// TIA Portal project "e009004v440" (V15.1) (continued)
   40: 'Reserva', class Reserva, trigger "DB_OP.DEF03" bit 15
   87: 'Falla al cerrar pinza posicionadora: Comprobar Sensores 29S4 y 29S5 + Electroválvula 43Y8 / FORMAGE : DEF MOUVEMENT FERMETURE PINCE 43Y8 : vérifier 29S4 29S5', class Fallos Pinza, trigger "DB_OP.DEF06" bit 14
   19: 'Falla térmica en freno de motor ajuste de ancho en etapa de Formado: Comprobar estado de Guardamotor Q09 / DF_QF9_1', class Fallos Formado, trigger "DB_OP.DEF02" bit 10
   68: 'Falla al subir araña: Comprobar sensores 25S7 y 25S8, y electroválvula 41Y3 / Falla al subir Araña: Comprobar Sensores 25S7 y 25S8 + Electroválvula 41Y3 / PREHENSEUR : DEF MOUVEMENT MONTEE 41Y3 : vérifier 25S7 25S8', class Fallos Araña, trigger "DB_OP.DEF05" bit 11
   71: 'Reserva', class Reserva, trigger "DB_OP.DEF05" bit 14
   21: 'Falla de excursión en Ajuste de ancho de Perfiladores: Comprobar 29S6, 29S7 + Encóder correspondiente / DEFAUT MOP PROFILEUSE : vérifier 29S6 29S7 ou codeur DP15', class Fallos Perfiladores, trigger "DB_OP.DEF02" bit 12
   67: 'Falla al bajar Araña: Comprobar Sensores 25S7 y 25S8 + Electroválvula 41Y2 / PREHENSEUR : DEF MOUVEMENT DESCENTE 41Y2 : vérifier 25S7 25S8', class Fallos Araña, trigger "DB_OP.DEF05" bit 10
   5: 'Falla en Variador Transporte Rolos: Comprobar estado de Variador VAR03 / Variateur OK Convoyeur Magasin', class Fallos Rolos, trigger "DB_OP.DEF01" bit 12
   24: 'Reserva', class Reserva, trigger "DB_OP.DEF02" bit 15
   95: 'Incoherencia en lectura de sensores 26S6 (Araña Arriba) y 26S7 (Araña Abajo) Soluciones Posibles: - Revise que el estado de ambos sensores sea correcto. - Revise el cableado de ambos sensores y asegúrese de que las señales llegan al panel observando los estados de los mismos desde el esquemático del PANEL / Falla al avanzar intercambiador de Almacenes: Comprobar Sensores 26S6 y 26S7 + Contactor KM01.1 / CHARGEMENT : DEF MOUVEMENT AVANCE MAGASIN : vérifier 26S6 26S7', class Fallos Almacenes, trigger "DB_OP.DEF06" bit 6
   101: 'Falla al subir Herramienta de Formado: Comprobar Sensores 28S5 y 28S6 + Relé 43K4 / FORMAGE : DEF MOUVEMENT MONTEE OUTIL 43K4 : vérifier 28S5 28S6', class Fallos Formado, trigger "DB_OP.DEF07" bit 12
   20: 'Falla en presión hidráulica en freno Perfiladores: Comprobar Sensor 23S4 / DEFAUT PRESSION HYDRAULIQUE FREIN PROFILEUSE : Vérifier 23S4', class Fallos Perfiladores, trigger "DB_OP.DEF02" bit 11
   50: 'Falla en Plegador 1 al intentar realizar plegado: Comprobar Sensores 31S7 y 31S8 + Relé 45K5 / PLIEUSE 1 : DEF MOUVEMENT AVANCE PLIAGE 45K5 : vérifier 31S7 et 31S8', class Fallos Plegadora, trigger "DB_OP.DEF04" bit 9
   111: 'Reserva', class Reserva, trigger "DB_OP.DEF07" bit 6
   65: 'Falla al transladar Araña (Avance): Comprobar Sensores 26S2 y 26S3 + Contactor KM02.1 / PREHENSEUR : DEF MOUVEMENT AVANCE KM02_1 : vérifier 26S2 26S3', class Fallos Araña, trigger "DB_OP.DEF05" bit 8
   53: 'Falla en Plegador 2 al intentar activar fijación: Comprobar Sensores 35S1 y 35S2 + Relé 47K1 / PLIEUSE 1 : DEF MOUVEMENT AVANCE BRIDAGE 45K3 : vérifier 31S5 et 31S6', class Fallos Plegadora, trigger "DB_OP.DEF04" bit 12
   109: 'Reserva', class Reserva, trigger "DB_OP.DEF07" bit 4
   39: 'Reserva', class Reserva, trigger "DB_OP.DEF03" bit 14
   56: 'Falla en Plegador 2 al intentar bajar primera extensión de prensa: Comprobar Sensores 35S7 y 35S8 + Relé 46K7 / PLIEUSE 2 : DEF MOUVEMENT AVANCE V2 47K7 : vérifier 35S7 et 35S8', class Fallos Plegadora, trigger "DB_OP.DEF04" bit 15
   54: 'Falla en Plegador 2 al intentar realizar plegado: Comprobar Sensores 35S3 y 35S4 + Relé 47K3 / PLIEUSE 1 : DEF MOUVEMENT AVANCE PLIAGE 45K5 : vérifier 31S7 et 31S8', class Fallos Plegadora, trigger "DB_OP.DEF04" bit 13
   108: 'Reserva', class Reserva, trigger "DB_OP.DEF07" bit 3
   86: 'Falla al bajar Bloqueador de Avance en etapa formador: Comprobar Sensores 29S1 y 29S2 + Electroválvula 43Y5 / FORMAGE : DEF MOUVEMENT DESCENTE BUTEE 43Y5 : vérifier 29S1 29S2', class Fallos Formado, trigger "DB_OP.DEF06" bit 13
   93: 'Falla al bajar Herramienta de Formado: Comprobar Sensores 28S5 y 28S6 + Relé 43K3 / FORMAGE : DEF MOUVEMENT DESCENTE OUTIL 43K3 : vérifier 28S5 28S6', class Fallos Formado, trigger "DB_OP.DEF06" bit 4
   34: 'Falla al bajar pinza en Plegadora: Comprobar Sensores 30S3 y 30S4 + Electroválvula 44Y3 / PLIEUSE : DEF MOUVEMENT DESCENTE PINCE 44Y3 : vérifier 30S3 et 30S4', class Fallos Plegadora, trigger "DB_OP.DEF03" bit 9
   27: 'Falla presión de Aire: Comprobar estado del Presostato 23S7 / DEFAUT AIR', class Fallos Generales, trigger "DB_OP.DEF02" bit 2
   115: 'Reserva', class Reserva, trigger "DB_OP.DEF08" bit 10
   97: 'Falla al retroceder martillo de herramienta 1 en Formador: Comprobar Sensores 27S5 y 27S6 + Relé 42K4 / FORMAGE : DEF MOUVEMENT RECUL MARTEAU OUTIL 1 42K4 : vérifier 27S5 27S6', class Fallos Formado, trigger "DB_OP.DEF07" bit 8
   88: 'Reserva', class Reserva, trigger "DB_OP.DEF06" bit 15
   57: 'Falla en Plegador 1 al intentar desactivar fijación: Comprobar Sensores 31S5 y 31S6 + Relé 45K4 / PLIEUSE 1 : DEF MOUVEMENT RECUL BRIDAGE 45K4 : vérifier 31S5 et 31S6', class Fallos Plegadora, trigger "DB_OP.DEF04" bit 0
   26: 'Falla de seguridad: Comprobar seguridades y relé de seguridad KAU1 / ATTENTE MISE EN SERVICE', class Fallos Generales, trigger "DB_OP.DEF02" bit 1
   18: 'Falla térmica en motor grupo hidráulico Plegadora: Comprobar estado de Guardamotor QM013.1 / DF_QM013_1 PLIEUSE : Moteur Groupe HYdraulique', class Fallos Plegadora, trigger "DB_OP.DEF02" bit 9
   36: 'Falla al activar alineacion X de Pieza en Plegadora: Comprobar Sensores 21S5, 21S6, 36S1 y 36S2 + Relé 46K5 / PLIEUSE : DEF MOUVEMENT TAQUAGE X 46K5 : vérifier 21S5 21S6 36S1 36S2', class Fallos Plegadora, trigger "DB_OP.DEF03" bit 11
   7: 'Falla en etapa de Potencia de variadores Perfiladores: Comprobar el estado de U13.2, U13.9, U13.12, U13.15 y U13.17 en Tablero T02 / DF_QM04 PROFILEUSE : Moteur 1,2,3 ou 4', class Fallos Perfiladores, trigger "DB_OP.DEF01" bit 14
   25: 'Falla alimentación de Entradas: Comprrobar estado de Térmica Q6 / ATTENTE MISE SOUS TENSION', class Fallos Generales, trigger "DB_OP.DEF02" bit 0
   104: 'Reserva', class Reserva, trigger "DB_OP.DEF07" bit 0
   96: 'Reserva', class Reserva, trigger "DB_OP.DEF06" bit 7
   77: 'Falla en Plegador 1 al intentar subir segunda extensión de prensa: Comprobar Sensores 32S5 y 32S6 + Relé 46K3 / PLIEUSE 1 : DEF MOUVEMENT AVANCE V3 46K3 : vérifier 32S5 32S6', class Fallos Plegadora, trigger "DB_OP.DEF05" bit 4
   8: 'Falla presente en CU Plegadores: Compruebe estado de CPU10', class Fallos Plegadora, trigger "DB_OP.DEF01" bit 15
   78: 'Falla en Plegador 2 al intentar subir segunda extensión de prensa: Comprobar Sensores 35S7 y 35S8 + Relé 48K1 / PLIEUSE 1 : DEF MOUVEMENT AVANCE V3 46K3 : vérifier 32S5 32S6', class Fallos Plegadora, trigger "DB_OP.DEF05" bit 5
   17: 'Falla límite de Seguridad en Plegador 2: Compruebe Sensor límite de carrera correspondiente / DF_VAR12 :PLIEUSE 2 : ServoVariateur OK', class Fallos Plegadora, trigger "DB_OP.DEF02" bit 8
   75: 'Reserva', class Reserva, trigger "DB_OP.DEF05" bit 2
   106: 'Reserva', class Reserva, trigger "DB_OP.DEF07" bit 1
   1: 'Falla térmica en motor refrigeración de grupo hidráulico Plegadora: Comprobar estado de Guardamotor QM013.2 / Moteur OK refroidisseur GH plieuse', class Fallos Perfiladores, trigger "DB_OP.DEF01" bit 8
   9: 'Falla de seguridad presente en CU Plegadores: Compruebe estado de CPU10', class Fallos Plegadora, trigger "DB_OP.DEF01" bit 0
   84: 'Reserva', class Reserva, trigger "DB_OP.DEF06" bit 11
   98: 'Falla al retroceder matriz de herramienta 1 en Formador: Comprobar Sensores 27S7 y 27S8 + Relé 42K6 / FORMAGE : DEF MOUVEMENT RECUL MATRICE OUTIL 1 42K6 : vérifier 27S7 27S8', class Fallos Formado, trigger "DB_OP.DEF07" bit 9
   92: 'Falla al avanzar matriz de herramienta 2 en Formador: Comprobar Sensores 28S3 y 28S4 + Relé 43K1 / FORMAGE : DEF MOUVEMENT AVANCE MATRICE OUTIL 2 43K1 : vérifier 28S3 28S4', class Fallos Formado, trigger "DB_OP.DEF06" bit 3
   99: 'Falla al retroceder martillo de herramienta 1 en Formador: Comprobar Sensores 28S1 y 28S2 + Relé 42K8 / FORMAGE : DEF MOUVEMENT RECUL MARTEAU OUTIL 2 42K8 : vérifier 28S1 28S2', class Fallos Formado, trigger "DB_OP.DEF07" bit 10
   120: 'Reserva', class Reserva, trigger "DB_OP.DEF08" bit 15
   16: 'Falla límite de Seguridad en Plegador 1: Compruebe Sensor límite de carrera correspondiente', class Fallos Plegadora, trigger "DB_OP.DEF01" bit 7
   59: 'Falla en Plegador 1 al intentar subir prensa: Comprobar Sensores 32S1 y 32S2 + Relé 45K8 / PLIEUSE 1 : DEF MOUVEMENT RECUL V1 45K8 : vérifier 32S1 et 32S2', class Fallos Plegadora, trigger "DB_OP.DEF04" bit 2
   42: 'Falla al subir pinza en Plegadora: Comprobar Sensores 30S3 y 30S4 + Electroválvula 44Y4 / PLIEUSE : DEF MOUVEMENT MONTEE PINCE 44Y4 : vérifier 30S3 et 30S4', class Fallos Plegadora, trigger "DB_OP.DEF03" bit 1
   11: 'Falla térmica en grupo hidraulico de freno Perfiladores: Comprobar estado de Guardamotor QM06 / DF_QM06 : PROFILEUSE : GH frein OK', class Fallos Perfiladores, trigger "DB_OP.DEF01" bit 2
   102: 'Falla al retroceder Descargador: Comprobar Sensores 31S2 y 31S3 + Relé 45K2 / DECHARGEMENT : DEF RECUL ESCAMOTEUR 45K2 : vérifier 31S2 31S3', class Fallos Descargador, trigger "DB_OP.DEF07" bit 13
   52: 'Falla en Plegador 1 al intentar subir primera extensión de prensa: Comprobar Sensores 32S3 y 32S4 + Relé 46K1', class Fallos Plegadora, trigger "DB_OP.DEF04" bit 11
   76: 'Reserva', class Reserva, trigger "DB_OP.DEF05" bit 3
   81: 'Falla al avanzar ajuste de formado: Comprobar Contactor KM09.1 + Encóder correspondiente / FORMAGE : DEF MOUVEMENT AVANCE MOP KM09_1 : vérifier codeur 2', class Fallos Cinta, trigger "DB_OP.DEF06" bit 8
   107: 'Reserva', class Reserva, trigger "DB_OP.DEF07" bit 2
   15: 'Falla Rectificador de variadores Plegadores: Comprobar estado de AL10', class Fallos Plegadora, trigger "DB_OP.DEF01" bit 6
   80: 'Falla en Plegador 2 al intentar bajar segunda extensión de prensa: Comprobar Sensores 35S7 y 35S8 + Relé 48K2 / PLIEUSE 1 : DEF MOUVEMENT AVANCE V3 46K3 : vérifier 32S5 32S6', class Fallos Plegadora, trigger "DB_OP.DEF05" bit 7
   47: 'Reserva', class Reserva, trigger "DB_OP.DEF03" bit 6
   43: 'Falla al cerrar pinza en Plegadora: Comprobar Sensores 30S5 y 30S6 + Electroválvula 44Y6 / PLIEUSE : DEF MOUVEMENT FERMETURE PINCE 44Y6 : vérifier 30S5 et 30S6', class Fallos Plegadora, trigger "DB_OP.DEF03" bit 2
   13: 'Falla en Variador Transporte Cinta: Comprobar estado de VAR08 / DF_VAR08 : CONVOYEUR 2 : Variateur OK', class Fallos Cinta, trigger "DB_OP.DEF01" bit 4
   45: 'Falla al desactivar alineacion Y de Pieza en Plegadora: Comprobar Sensores 23S6 y 36S4 + Relé 46K6', class Fallos Plegadora, trigger "DB_OP.DEF03" bit 4
   105: 'Reserva', class Reserva, trigger "DB_OP.DEF07" bit 15
   38: 'Falla al desactivar alineacion Y de Pieza en Plegadora: Comprobar Sensores 23S5, 23S6, 36S3 y 36S4 + Relé 46K6', class Fallos Plegadora, trigger "DB_OP.DEF03" bit 13
   31: 'Falla de Atasco de pieza en Perfilador: Compobar Sensores 36S13, 36S14, 36S15 y 36S16 / DEFAUT BOURRAGE PROFILEUSE', class Fallos Perfiladores, trigger "DB_OP.DEF02" bit 6
   72: 'Reserva', class Reserva, trigger "DB_OP.DEF05" bit 15
   89: 'Falla al avanzar martillo de herramienta 1 en Formador: Comprobar Sensores 27S5 y 27S6 + Relé 42K3 / FORMAGE : DEF MOUVEMENT AVANCE MARTEAU OUTIL 1 42K3 : vérifier 27S5 27S6', class Fallos Formado, trigger "DB_OP.DEF06" bit 0
   114: 'Reserva', class Reserva, trigger "DB_OP.DEF08" bit 9
   10: 'Falla térmica en bomba de lubricación de Perfiladores: Comprobar estado de Guardamotor QM05 / DF_QM05 : PROFILEUSE :Pompes lubrifications OK', class Fallos Perfiladores, trigger "DB_OP.DEF01" bit 1
   4: 'Falla en Variador Transporte de Araña: Comprobar estado de Variador VAR02 / Variateur OK Axe Prehenseur', class Fallos Araña, trigger "DB_OP.DEF01" bit 11
   110: 'Reserva', class Reserva, trigger "DB_OP.DEF07" bit 5
   73: 'Falla al transladar Araña (Retroceder): Comprobar Sensores 26S2 y 26S3, y Contactor KM02.2 / PREHENSEUR : DEF MOUVEMENT RECUL KM02_2 : vérifier 26S2 26S3', class Fallos Araña, trigger "DB_OP.DEF05" bit 0
   44: 'Falla al desactivar alineacion X de Pieza en Plegadora: Comprobar Sensores 36S2 y 21S6 + Relé 46K5 / PLIEUSE : DEF MOUVEMENT TAQUAGE X 46K5 : vérifier 21S5 21S6 36S1 36S2', class Fallos Plegadora, trigger "DB_OP.DEF03" bit 3
   118: 'Reserva', class Reserva, trigger "DB_OP.DEF08" bit 13
   94: 'Falla al avanzar Descargador: Comprobar Sensores 31S2 y 31S3 + Relé 45K1 / DECHARGEMENT : DEF AVANCE ESCAMOTEUR 45K1 : vérifier 31S2 31S3', class Fallos Descargador, trigger "DB_OP.DEF06" bit 5
   58: 'Falla en Plegador 1 al intentar desactivar orden de plegado: Comprobar Sensores 31S7 y 31S8 + Relé 45K6 / PLIEUSE 1 : DEF MOUVEMENT RECUL PLIAGE 45K6 : vérifier 31S7 et 31S8', class Fallos Plegadora, trigger "DB_OP.DEF04" bit 1
   63: 'Falla en Plegador 2 al intentar subir prensa: Comprobar Sensores 35S5 y 35S6 + Relé 47K6 / PLIEUSE 1 : DEF MOUVEMENT RECUL V1 45K8 : vérifier 32S1 et 32S2', class Fallos Plegadora, trigger "DB_OP.DEF04" bit 6
   119: 'Reserva', class Reserva, trigger "DB_OP.DEF08" bit 14
   60: 'Falla en Plegador 1 al intentar bajar primera extensión de prensa: Comprobar Sensores 32S3 y 32S4 + Relé 46K2', class Fallos Plegadora, trigger "DB_OP.DEF04" bit 3
   23: 'Falla Seguridad de Perímetro: Comprobar Seguridad de puertas y tablero CPI / DF_RES01', class Fallos Generales, trigger "DB_OP.DEF02" bit 14
   32: 'Reserva / DF_RES01', class Reserva, trigger "DB_OP.DEF02" bit 7
   22: 'Falla de excursión en Ajuste de ancho de Formado: Comprobar 28S7, 28S8 + Encóder correspondiente / DEFAUT MOP CONVOYEUR2 : vérifier 28S7 28S8 ou codeur DP16', class Fallos Formado, trigger "DB_OP.DEF02" bit 13
   79: 'Falla en Plegador 1 al intentar bajar segunda extensión de prensa: Comprobar Sensores 32S5 y 32S6 + Relé 46K3 / PLIEUSE 2 : DEF MOUVEMENT AVANCE V3 48K1 : vérifier 36S7 36S8', class Fallos Plegadora, trigger "DB_OP.DEF05" bit 6

text list "SelecciónPlegadora": 0 'Sin selección'; 1 'Plegador 1'; 2 'Plegador 2'; 3 'Tenaza'

text list "Modo": 0 'Detenido / ARRET'; 1 'Modo Manual / MANUEL'; 2 'Modo Automático / AUTO'; 3 'En Ciclo / CYCLE'; 4 'Finalizando Ciclo / FIN CYCLE'

text list "RC1": 0 '00: Sin selección / 00: ACQUITTEMENT'; 1 '01: Intercambiador de almacenes - Avance / 01 : Avance Magasin (mag 1)'; 2 '02: Intercambiador de almacenes - Retroceso / 02 : Recul Magasin (mag 2)'; 11 '11: Transporte Araña - Avance / 11 : Préhenseur Avance'; 12 '12: Transporte Araña - Retroceso / 12 : Préhenseur Recul'; 13 '13: Araña - Bajar sobre Almacén 1 / 13 : Préhenseur Magasin 1'; 14 '14: Araña - Bajar sobre Almacén 2 / 14 : Préhenseur Magasin 2'; 15 '15: Araña - Bajar / 15 : Préhenseur Descente'; 16 '16: Araña - Subir / 16 : Préhenseur Montée'; 20 '20: Tulipas de Araña - Aire en todas ON / 20 :Flambage 1 à 3 Avance'; 21 '21: Tulipas de Araña - Aire en todas OFF / 21: Flambage 1 à 3 Recul'; 22 '22: Tulipas de Araña - Aire en Grupo 1 ON / 22 : Flambage 1 Avance'; 23 '23: Tulipas de Araña - Aire en Grupo 1 OFF / 23 : Flambage 1 Recul'; 24 '24: Tulipas de Araña - Aire en Grupo 2 ON / 24 : Flambage 2 Avance'; 25 '25: Tulipas de Araña - Aire en Grupo 2 OFF / 25 : Flambage 2 Recul'; 26 '26: Tulipas de Araña - Aire en Grupo 3 ON / 26 : Flambage 3 Avance'; 27 '27: Tulipas de Araña - Aire en Grupo 3 OFF / 27 : Flambage 3 Recul'; 30 '30: Tulipas de Araña - Vacío en Todas ON / 30 :Aspiration 1 à 3 Avance'; 31 '31: Tulipas de Araña - Vacío en Todas OFF / 31: Aspiration 1 à 3 Recul'; 32 '32: Tulipas de Araña - Vacío en Grupo 1 ON / 32 : Aspiration 1 Avance'; 33 '33: Tulipas de Araña - Vacío en Grupo 1 OFF / 33 : Aspiration 1 Recul'; 34 '34 : Tulipas de Araña - Vacío en Grupo 2 ON / 34 : Aspiration 2 Avance'; 35 '35: Tulipas de Araña - Vacío en Grupo 2 OFF / 35 : Aspiration 2 Recul'; 36 '36: Tulipas de Araña - Vacío en Grupo 3 ON / 36 : Aspiration 3 Avance'; 37 '37: Tulipas de Araña - Vacío en Grupo 3 OFF / 37 : Aspiration 3 Recul'; 41 '41: Transporte Rolos - Avance / 41 avance Convoyeur 1'; 42 '42: Transporte Rolos - Retroceso / 42 Recul Convoyeur 1'; 51 '51: Ajuste de profundidad Perfiladores - Hacia Consigna / 51 : MOP Profileuse Consigne'; 52 '52: Ajuste de profundidad Perfiladores - Cerrar / 52 : Avance MOP Profileuse'; 53 '53: Ajuste de profundidad Perfiladores - Abrir / 53 : Recul MOP Profileuse'; 54 '54: Ajuste de profundidad Perfiladores - Freno / 54 : Frein MOP profileuse'; 55 '55: Perfiladores - Retroceso / 55 : Avance Profileuse'; 56 '56: Perfiladores - Avance / 56 : Recul Profileuse'

text list "RC2": 0 '00: Sin Selección / 00: ACQUITTEMENT'; 1 '01: Plegadora - Avance Tenaza / 01:Pince: Avance'; 2 '02: Plegadora - Retroceso Tenaza / 02:Pince: Recul'; 3 '03: Plegadora - Bajar Tenaza / 03:Pince: Descente'; 4 '04: Plegadora - Subir Tenaza / 04:Pince: Montée'; 5 '05: Plegadora - Abrir Tenaza / 05:Pince: ouverture'; 6 '06: Plegadora - Cerrar Tenaza / 06:Pince: Fermeture'; 7 '07: Plegadora - Alineación X / 07:taquage X'; 8 '08: Plegadora - Alineación Y / 08:taquage Y'; 9 '09: Plegadora - Subir Cepillos / 09: brosse'; 10 '10: Plegador 1 - Bloquear Prensa / 10:PLIEUSE 1: bridage Avance'; 11 '11: Plegador 1 - Desbloquear Prensa / 11:PLIEUSE 1: bridage Recul'; 12 '12: Plegador 1 - Bajar Prensa / 12:PLIEUSE 1: V1 Avance'; 13 '13: Plegador 1 - Subir Prensa / 13:PLIEUSE 1: V1 Recul'; 14 '14: Plegador 1 - Bajar Extension Prensa 1 / 14:PLIEUSE 1: V2 Avance'; 15 '15: Plegador 1 - Subir Extension Prensa 1 / 15:PLIEUSE 1: V2 Recul'; 16 '16: Plegador 1 - Bajar Extension Prensa 2 / 16:PLIEUSE 1: V3 Avance'; 17 '17: Plegador 1 - Subir Extension Prensa 2 / 17:PLIEUSE 1: V3 Recul'; 18 '18: Plegador 1 - Subir / 18:PLIEUSE 1: Montée'; 19 '19: Plegador 1 - Bajar / 19:PLIEUSE 1: Descente'; 20 '20: Plegador 2 - Bloquear Prensa / 20:PLIEUSE 2: bridage Avance'; 21 '21: Plegador 2 - Desbloquear Prensa / 21:PLIEUSE 2: bridage Recul'; 22 '22: Plegador 2 - Bajar Prensa / 22:PLIEUSE 2: V1 Avance'; 23 '23: Plegador 2 - Subir Prensa / 23:PLIEUSE 2: V1 Recul'; 24 '24: Plegador 2 - Bajar Extension Prensa 1 / 22:PLIEUSE 2: V1 Avance'; 25 '25: Plegador 2 - Subir Extension Prensa 1 / 23:PLIEUSE 2: V1 Recul'; 26 '26: Plegador 2 - Bajar Extension Prensa 2 / 26:PLIEUSE 2: V3 Avance'; 27 '27: Plegador 2 - Subir Extension Prensa 2 / 27:PLIEUSE 2: V3 Recul'; 28 '28: Plegador 2 - Subir / 28:PLIEUSE 2: Montée'; 29 '29: Plegador 2 - Bajar / 29:PLIEUSE 2: Descente'; 31 '31: Pinza - Avance / 31 : Avance Pince'; 32 '32: Pinza - Retroceso / 32 : Recul Pince'; 33 '33: Pinza - Abrir / 33: Ouverture Pince'; 34 '34: Pinza - Cerrar / 34: Fermeture Pince'; 35 '35: Formador - Subir Tope / 35: Montée Butée'; 36 '36: Formador - Bajar Tope / 36: Descente Butée'; 37 '37: Formador - Ajuste de profundidad - Hacia Consigna / 37: Position Consigne'; 38 '38: Formador - Ajuste de profundidad - Avance / 38: Rapproche ( - )'; 39 '39: Formador - Ajuste de profundidad - Retroceso / 39: Ecartement ( + )'; 40 '40: Formador - Bajar Herramientas / 40: Descente Ensemble'; 41 '41: Formador - Subir Herramientas / 41: Montée Ensemble'; 42 '42: Formador - Herramienta 1 - Martillo ON / 42: MARTEAU : Avance Outil 1'; 43 '43: Formador - Herramienta 1 - Martillo OFF / 43: MARTEAU : Recul Outil 1'; 44 '44: Formador - Herramienta 1 - Matriz ON / 44: MATRICE : Avance Outil 1'; 45 '45: Formador - Herramienta 1 - Matriz OFF / 45: MATRICE : Recul Outil 1'; 46 '46: Formador - Herramienta 2 - Martillo ON / 46: MARTEAU : Avance Outil 2'; 47 '47: Formador - Herramienta 2 - Martillo OFF / 47: MARTEAU : Recul Outil 2'; 48 '48: Formador - Herramienta 2 - Matriz ON / 48: MATRICE : Avance Outil 2'; 49 '49: Formador - Herramienta 2 - Matriz OFF / 49: MATRICE : Recul Outil 2'; 61 '61: Plegador 1 - Avance (apertura) / 61: PLIEUSE 1 : Ecartement +'; 62 '62: Plegador 1 - Retroceso (cierre) / 62: PLIEUSE 1 : Rapproche -'; 65 '65: Plegador 2 - Avance (apertura) / 65: PLIEUSE 2 : Ecartement +'; 66 '66: Plegador 2 - Retroceso (cierre) / 66: PLIEUSE 2 : Rapproche -'; 70 '70: Descargador - Avance / 70: Avance Escamoteur'; 71 '71: Descargador - Retroceso / 71: Recul Escamoteur'; 91 '91: Transporte Cinta - Avance / 91: Avance Convoyeur 2'; 92 '92: Transporte Cinta - Retroceso / 92: Recul Convoyeur 2'

text list "Warnings": 0 'Sin Warnings'; 1 'Reconocimiento de Fallas solo es posible en Modo Manual'; 2 'No es posible intercambiar almacenes si la Araña no está completamente arriba'; 4 ''; 8 'Los plegadores no pueden desplazarse si sus prensas no estan completamente abiertas'; 16 'Los plegados solo son posibles con las prensas abajo'; 32 'Para poder bloquear los plegadores es becesario que las prensas estén abajo'; 64 'Solo es posible accionar las herramientas si el formador está abajo'; 128 ''; 254 ''; 512 ''; 1024 ''; 2048 ''; 4096 ''

text list "Estados_PL": 0 'Detenido'; 512 'Esperando Pieza'; 1024 'Ingresando Pieza'; 2048 'Posicionando Plegadores para Primer Plegado'; 4096 'Realizando Primer Plegado'; 8192 'Realizando Segundo Plegado'; 16384 'Entregando Pieza'; 2 'Alineando Pieza'; 4 'Posicionando Plegadores para Segundo Plegado'; 8 'Posicionando Plegadores para Entrega de Pieza'; 16 'Posicionando Plegadores para Espera'

text list "Estados_F": 128 'Detenido'; 512 'Esperando'; 1024 'Formando Pieza en Esquina 1 con Herramienta 1'; 2048 'Formando Pieza en Esquina 1 con Herramienta 2'; 4096 'Formando Pieza en Esquina 2 con Herramienta 1'; 8192 'Formando Pieza en Esquina 2 con Herramienta 2'; 16384 'Entregando Pieza'; -32768 'Posicionando Pieza en Esquina 1 con Herramienta 1'; 1 'Posicionando Pieza en Esquina 1 con Herramienta 2'; 2 'Posicionando Pieza en Esquina 2 con Herramienta 1'; 4 'Posicionando Pieza en Esquina 2 con Herramienta 2'; 8 'Posicionando Pieza para Entrega'; 16 'Posicionando Pinza para Recepción de Pieza'

text list "Transiciones_PL": 0 'Condición de avance: Sin pieza en Plegadora'; 16 'Condición de avance: Posición de Espera alcanzada'; 512 'Condición de avance: Nueva Pieza en Plegadora'; 2 'Condición de avance: Alineadores Activos'; 2048 'Condición de avance: Posición de Plegado de Patas alcanzada'; 4 'Condición de avance: Posición de Plegado de Techo alcanzada'; 8 'Condición de avance: Posición de Entrega alcanzada'; 1024 'Condición de avance: Tenaza Plegadora adentro (Abierta)'; 4096 'Condición de avance: Plegado de Patas Activo'; 8192 'Condición de avance: Plegado de Techo Activo'; 16384 'Condición de avance: Pieza entregada a Descargador'

text list "Transiciones_F": 128 'Condición de avance: Sin Pieza en Pinza'; 512 'Condición de avance: Nueva Pieza en Final de Cinta'; 1024 'Condición de avance: Formado con Herramienta 1 Listo'; 2048 'Condición de avance: Formado con Herramienta 2 Listo'; 4096 'Condición de avance: Formado con Herramienta 1 Listo'; 8192 'Condición de avance: Formado con Herramienta 2 Listo'; 16384 'Condición de avance: Pieza entregada a Plegadora'; -32768 'Condición de avance: Posición de E1H1 alcanzada'; 1 'Condición de avance: Posición de E1H2 alcanzada'; 2 'Condición de avance: Posición de E2H1 alcanzada'; 4 'Condición de avance: Posición de E2H2 alcanzada'; 8 'Condición de avance: Posición de Entrega alcanzada'; 16 'Condición de avance: Posición de Recepción alcanzada'

text list "Proveedor": 0 ''; 1 'A'; 2 'B'; 3 'C'; 4 'D'; 5 'E'; 6 'F'

graphic list "General - Araña": 0..1 'Araña 1 G'; 1 'Araña 2_1'

graphic list "General - Almacén": 0..1 'Almacen 1 G'; 1 'Almacen 2_1'

graphic list "General - Rolos": 0..1 'Rolos 1 G'; 1 'Rolos 2_3'

graphic list "General - Perfiladores": 0..1 'Perfiladores 1 G'; 1 'Perfiladores 2_1'

graphic list "General - Cinta": 0..1 'Cinta G'; 1 'Cinta 2_1'

graphic list "General - Pinza": 0..1 'Pinza G'; 1 'Pinza 2_1'

graphic list "General - Formador": 0..1 'F1_G'; 1 'F1R'

graphic list "General - Plegadora": 0..1 'Plegador 1 G'; 1 'Plegador 2_1'

graphic list "General - Descargador": 0..1 'Descargador G'; 1 'Descargador 2_1'

graphic list "Intercambiador": 0..1 'ALM 2_1'; 1 'ALM 1'

graphic list "Grupo 3 - Plegadora": 0 'Pleg'; 1 'Pleg2'

graphic list "Grupo 3 - Descargador": 0..1 'Desc G'; 1 'Desc2'

graphic list "Grupo 3 - Pinza1": 0..1 'P2_G'; 1 'P2R'

graphic list "Pleg3": 1 'PLEG3b'; 2..3 'pleg_1'

graphic list "Grupo 1 - Rolos": 1 'Rolos 2 G'; 1 'Rolos 2b'

graphic list "Grupo 1 - Araña": 1 'Araña3b'; 2..3 'Araña3 G'

graphic list "Grupo 1 - Almacén A": 1 'ALM 2 G'; 2..3 'ALM 1 G'

graphic list "Grupo 1 - Almacén B": 1 'ALM 2b'; 2..3 'ALM 1b_1'

graphic list "Grupo 2 - Perfilador": 1 'PERFIb'; 2..3 'PERFI G'

graphic list "Grupo 2 - Cinta": 1 'CINb'; 2..3 'CIN G'

graphic list "Grupo 2 - Formador": 1 'Piqb'; 2..3 'Piq_1'

graphic list "Formador": 1 'F1R'; 2..3 'F1_G'

graphic list "Araña": 1 'Araña4b'; 2..3 'Araña4C'

graphic list "Rolos": 1 'Rolos 3b'; 2..3 'Rolos 3 G'

graphic list "GeneralBase": 0 'Base G'; 1 'BaseRoja'

graphic list "Estado": 0 'PilotLight_Round_GN_Off_256c'; 1 'PilotLight_Round_GN_On_256c'

graphic list "CheckBox": 0 'outline_check_box_outline_blank_black_18dp'; 1 'outline_check_box_black_18dp'

graphic list "CheckBox_Neg": 1 'outline_check_box_outline_blank_black_18dp'; 0 'outline_check_box_black_18dp'

graphic list "Pleg3_1": 1 'PLEG3b'; 2..3 'PLEG3_1'

graphic list "Grupo 3 - Pinza1_1": 0..1 'P2'; 1 'P2R'

graphic list "Formador_1": 1 'F2R'; 2..3 'F2C'

graphic list "Formador_2": 1 'F2R'; 2..3 'F2C'

recipe "Pieza": A <- "Receta\Recetas.A", B <- "Receta\Recetas.B", C <- "Receta\Recetas.C", D <- "Receta\Recetas.D", F1 <- "Receta\Recetas.F1", F2 <- "Receta\Recetas.F2", F3 <- "Receta\Recetas.F3", F4 <- "Receta\Recetas.F4", PL1_1 <- "Receta\Recetas.PL1_1", PL1_2 <- "Receta\Recetas.PL1_2", PL2_1 <- "Receta\Recetas.PL2_1", PL2_2 <- "Receta\Recetas.PL2_2"

screen "HabAlarmas9" 1280x768, template "Template"
   TextField "Campo de texto_1" at 117,85 size 37x18; Text '113 -'
   TextField "Campo de texto_2" at 117,129 size 37x18; Text '114 -'
   TextField "Campo de texto_3" at 117,173 size 37x18; Text '115 -'
   TextField "Campo de texto_4" at 117,217 size 367x18; Text '116 - Inconsistencia de Presencia de pieza en Transporte de Rolos'
   TextField "Campo de texto_5" at 117,261 size 37x18; Text '117 -'
   TextField "Campo de texto_6d" at 117,305 size 37x18; Text '118 -'
   TextField "Campo de texto_7" at 117,349 size 37x32; Text '119 -'
   TextField "Campo de texto_8" at 117,393 size 37x32; Text '120 -'
   TextField "Campo de texto_9" at 117,437 size 342x18; Text '121 - Inconsistencia de Presencia de pieza en en Descargador'
   Switch "Interruptor_1" at 48,77 size 59x33; TextOff 'SI'; TextOn 'NO'; CaptionText 'Switch'; PictureOff "Check"; PictureOn "UnCheck"
      ProcessValue <- "Desactivar_Falla113"
   Switch "Interruptor_2" at 48,121 size 59x33; TextOff 'SI'; TextOn 'NO'; CaptionText 'Switch'; PictureOff "Check"; PictureOn "UnCheck"
      ProcessValue <- "Desactivar_Falla114"
   Switch "Interruptor_3" at 48,165 size 59x33; TextOff 'SI'; TextOn 'NO'; CaptionText 'Switch'; PictureOff "Check"; PictureOn "UnCheck"
      ProcessValue <- "Desactivar_Falla115"
   Switch "Interruptor_4" at 48,209 size 59x33; TextOff 'SI'; TextOn 'NO'; CaptionText 'Switch'; PictureOff "Check"; PictureOn "UnCheck"
      ProcessValue <- "Desactivar_Falla116"
   Switch "Interruptor_5" at 48,253 size 59x33; TextOff 'SI'; TextOn 'NO'; CaptionText 'Switch'; PictureOff "Check"; PictureOn "UnCheck"
      ProcessValue <- "Desactivar_Falla117"
   Switch "Interruptor_6" at 48,297 size 59x33; TextOff 'SI'; TextOn 'NO'; CaptionText 'Switch'; PictureOff "Check"; PictureOn "UnCheck"
      ProcessValue <- "Desactivar_Falla118"
   Switch "Interruptor_7" at 48,341 size 59x33; TextOff 'SI'; TextOn 'NO'; CaptionText 'Switch'; PictureOff "Check"; PictureOn "UnCheck"
      ProcessValue <- "Desactivar_Falla119"
   Switch "Interruptor_8" at 48,385 size 59x33; TextOff 'SI'; TextOn 'NO'; CaptionText 'Switch'; PictureOff "Check"; PictureOn "UnCheck"
      ProcessValue <- "Desactivar_Falla120"
   Switch "Interruptor_9" at 48,429 size 59x33; TextOff 'SI'; TextOn 'NO'; CaptionText 'Switch'; PictureOff "Check"; PictureOn "UnCheck"
      ProcessValue <- "Desactivar_Falla121"
   TextField "Campo de texto_15" at 38,32 size 262x22; Text 'Configuración de habilitación de Alarmas'
   Button "Botón_2" at 1010,33 size 51x51; TextOff '<'
      on Click: ActivateScreen("HabAlarmas7", 0)
   Button "Botón_3" at 1202,33 size 51x51; TextOff '>'
   Circle "Círculo_2" at 24,87 size 12x12
      Appearance <- "Alarma 1"
   Circle "Círculo_3" at 25,131 size 12x12
      Appearance <- "Alarma 114"
   Circle "Círculo_4" at 25,175 size 12x12
      Appearance <- "Alarma 115"
   Circle "Círculo_5" at 24,87 size 12x12
      Appearance <- "Alarma 113"
   Circle "Círculo_6" at 25,219 size 12x12
      Appearance <- "Alarma 116"
   Circle "Círculo_7" at 25,263 size 12x12
      Appearance <- "Alarma 117"
   Circle "Círculo_8" at 25,307 size 12x12
      Appearance <- "Alarma 118"
   Circle "Círculo_9" at 25,351 size 12x12
      Appearance <- "Alarma 119"
   Circle "Círculo_10" at 25,395 size 12x12
      Appearance <- "Alarma 120"
   Circle "Círculo_11" at 25,439 size 12x12
      Appearance <- "Alarma 121"
   Button "Template_Plantilla_Bouton_0" at 1085,715 size 193x53; TextOff 'ALARMAS / DEFAUT'
      on Press: ActivateScreen("eProC - Alarmas", 0)
   Button "Template_Plantilla_Bouton_2" at 1085,715 size 193x53; TextOff 'ALARMAS / DEFAUT'
      on Press: ActivateScreen("eProC - Alarmas", 0)
      Visibility <- "DB_OP.P_DEFAUT"
   Button "Template_Plantilla_Botón_3" at 1085,688 size 193x29; TextOff 'DESACT. TEMP. ALARMAS'

screen "eProC - Alarmas" 1280x768, template "Template"
   AlarmView "Vue des alarmes_1" at 13,32 size 1254x587; ColumnTextDate 'Fecha / Date'; ColumnTextDevice 'Control / Automate'; ColumnTextAckGroup 'GR'; ColumnTextNumber 'Nº / N°'; ColumnTextAlarmState 'Estado / Etat'; ColumnTextAlarmText 'Texto / Texte'; ColumnTextTime 'Hora / Heure'
   Button "Bouton" at 1084,638 size 195x53; TextOff 'RECONOCER ALARMAS / ACQUITEMENT'
      on Press: SetBit("DB_OP.ACQ_DEFAUT")
      Appearance <- "DB_OP.P_DEFAUT"
   Button "Botón_17" at 936,638 size 150x53; TextOff 'DESACT. TEMP. ALARMAS'; Authorization "Nivel 2"
      on Click: ActivateScreen("HabAlarmas1", 0)
   Button "Botón_1" at 788,638 size 150x53; TextOff 'HISTORIAL'
      on Click: ActivateScreen("eProC - Historal", 0)
   Button "Template_Plantilla_Bouton_0" at 1085,715 size 193x53; TextOff 'ALARMAS / DEFAUT'
      on Press: ActivateScreen("eProC - Alarmas", 0)
   Button "Template_Plantilla_Bouton_2" at 1085,715 size 193x53; TextOff 'ALARMAS / DEFAUT'
      on Press: ActivateScreen("eProC - Alarmas", 0)
      Visibility <- "DB_OP.P_DEFAUT"

